REGION Network 26: fermer cv01 en 4k
   #_w1 := "EtatMode4k" AND NOT "CV01_ManAuto";
   IF #_w1 THEN
       "unscal_ret_val" := UNSCALE(IN := 0.0,
                               HI_LIM := 100.0,
                               LO_LIM := 0.0,
                               BIPOLAR := "always_0",
                               OUT => "CMD_CV_01");
       "PLC_to_Epics".CV01.sSetVAuto := 0.0;
   END_IF;
END_REGION

REGION Network 27: 2K mode - close CV02 after precooling the 2K line
   #_w1 := "EtatMode2K" AND (#S8step > 4);
   IF #_w1 THEN
       "unscal_ret_val_1" := UNSCALE(IN := 0.0,
                               HI_LIM := 100.0,
                               LO_LIM := 0.0,
                               BIPOLAR := "always_0",
                               OUT => "CMD_CV_02");
       "PLC_to_Epics".CV02.sSetVAuto := 0.0;
   END_IF;
END_REGION

REGION Network 28: Init 2K mode
   #_w1 := "EtatMode2K" AND NOT "2KModeStart_mem";   // rising edge of "EtatMode2K"
   "2KModeStart_mem" := "EtatMode2K";
   IF #_w1 THEN
       #S8step := 4;
       "unscal_ret_val" := UNSCALE(IN := "S8_parameters".CV01_Init,
                               HI_LIM := 100.0,
                               LO_LIM := 0.0,
                               BIPOLAR := "always_0",
                               OUT => "CMD_CV_01");
       "PLC_to_Epics".CV01.sSetVAuto := "S8_parameters".CV01_Init;
   END_IF;
END_REGION

REGION Network 29: 2K mode - precooling (step4)
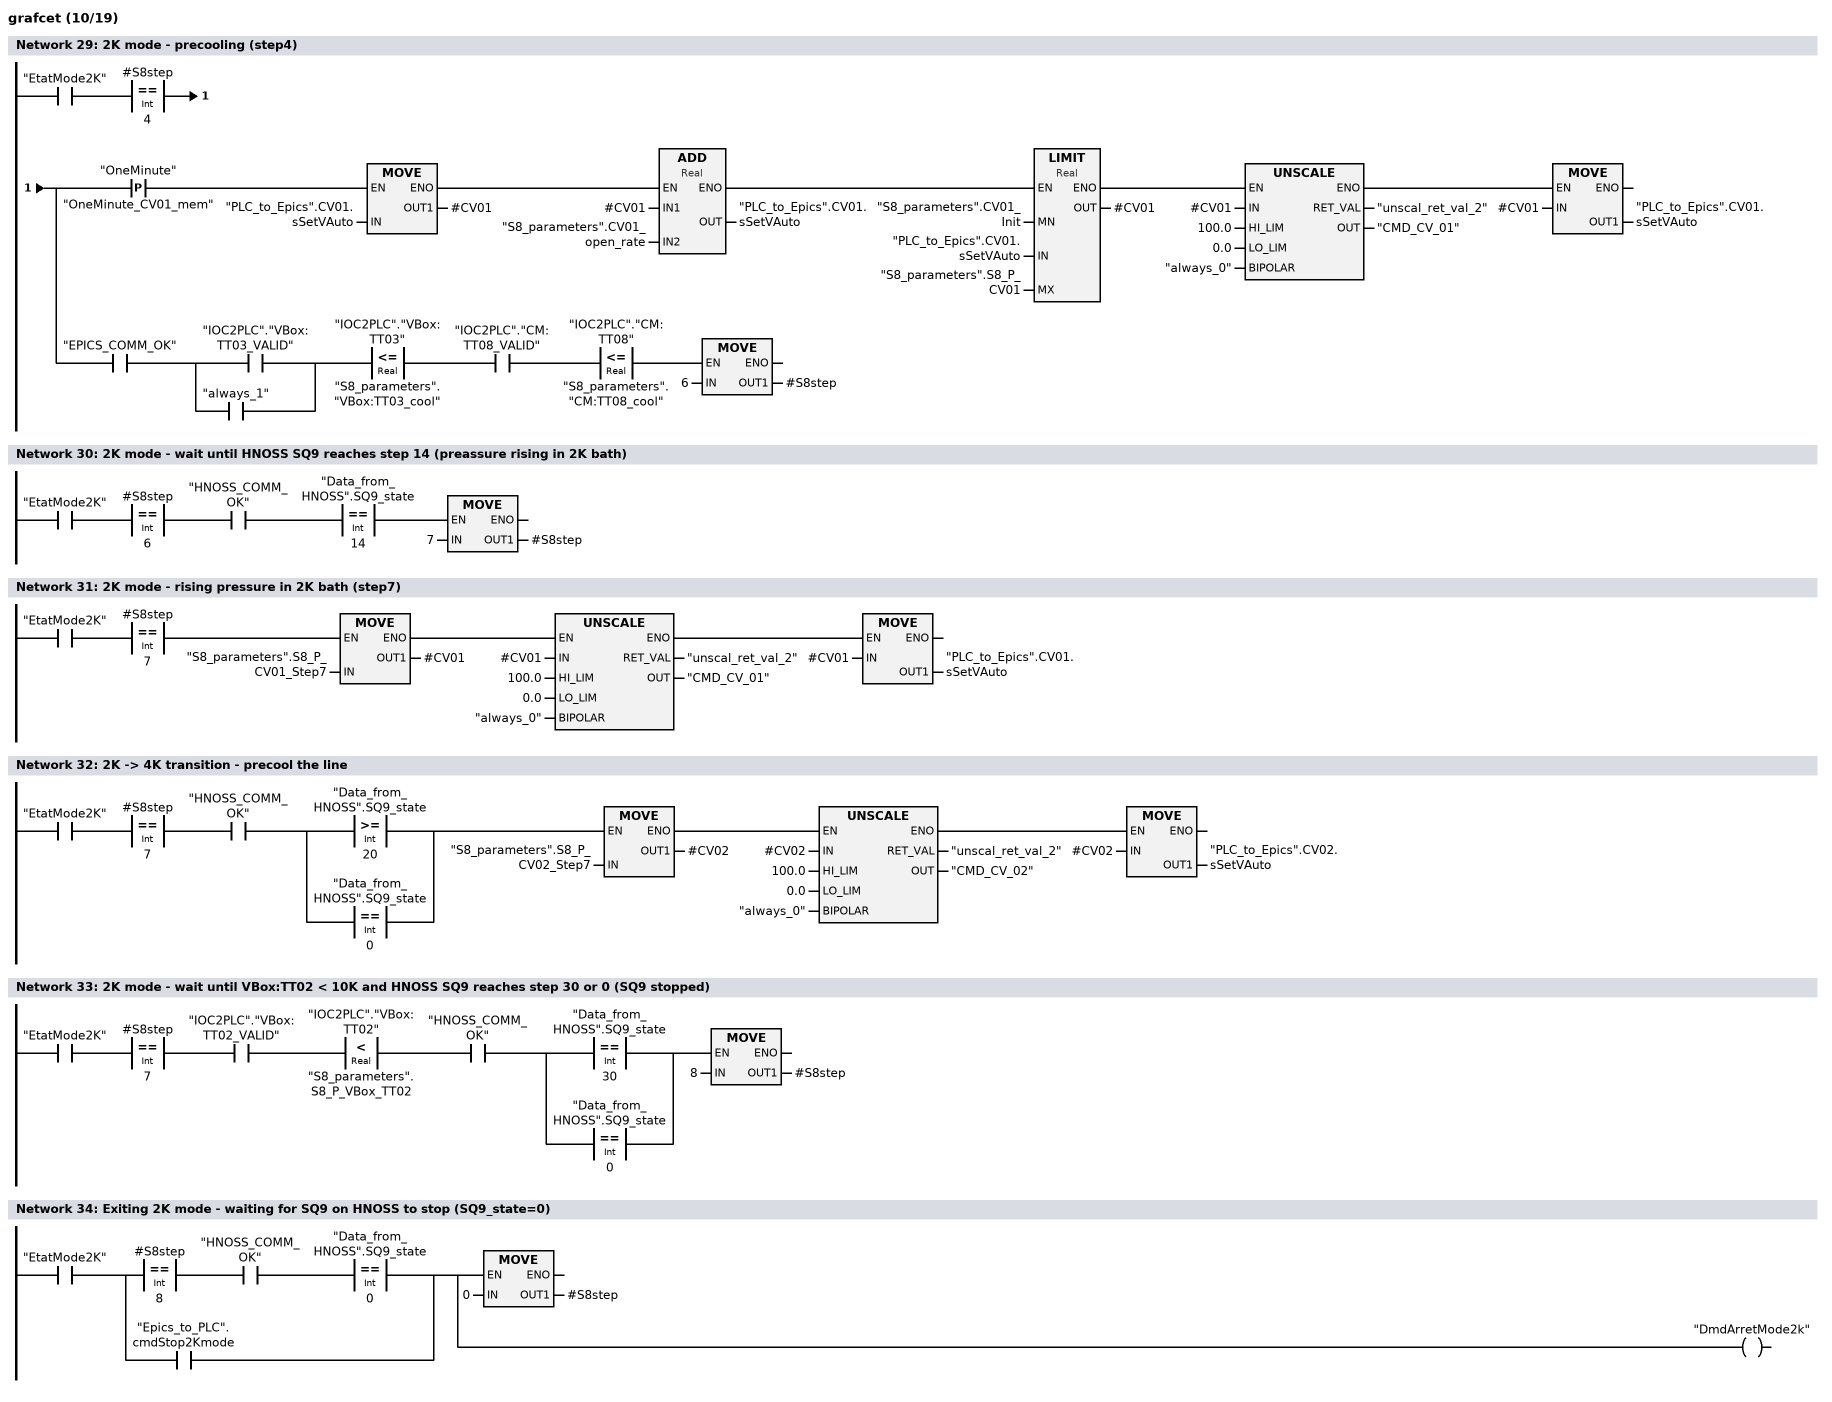
   // ENO of a box is taken as its EN; it also drops when the box reports an error
   #_w1 := "EtatMode2K" AND (#S8step = 4);
   #_w2 := #_w1 AND "OneMinute" AND NOT "OneMinute_CV01_mem";   // rising edge of "OneMinute"
   "OneMinute_CV01_mem" := "OneMinute";
   IF #_w2 THEN
       #CV01 := "PLC_to_Epics".CV01.sSetVAuto;
       "PLC_to_Epics".CV01.sSetVAuto := #CV01 + "S8_parameters".CV01_open_rate;
       #CV01 := LIMIT(MN := "S8_parameters".CV01_Init, IN := "PLC_to_Epics".CV01.sSetVAuto, MX := "S8_parameters".S8_P_CV01);
       "unscal_ret_val_2" := UNSCALE(IN := #CV01,
                               HI_LIM := 100.0,
                               LO_LIM := 0.0,
                               BIPOLAR := "always_0",
                               OUT => "CMD_CV_01");
       "PLC_to_Epics".CV01.sSetVAuto := #CV01;
   END_IF;
   IF #_w1 AND "EPICS_COMM_OK" AND ("IOC2PLC"."VBox:TT03_VALID" OR "always_1") AND ("IOC2PLC"."VBox:TT03" <= "S8_parameters"."VBox:TT03_cool") AND "IOC2PLC"."CM:TT08_VALID" AND ("IOC2PLC"."CM:TT08" <= "S8_parameters"."CM:TT08_cool") THEN
       #S8step := 6;
   END_IF;
END_REGION

REGION Network 30: 2K mode - wait until HNOSS SQ9 reaches step 14 (preassure rising in 2K bath)
   RUNG wire#powerrail
      Contact( "EtatMode2K" )
      { S7_Templates := "SrcType := Int" } EQ_Contact(in1 := #S8step, in2 := 6)
      Contact( "HNOSS_COMM_OK" )
      { S7_Templates := "SrcType := Int" } EQ_Contact(in1 := "Data_from_HNOSS".SQ9_state, in2 := 14)
      { S7_GenerateENO := "TRUE" } Move(in := 7, out1 => #S8step)
   END_RUNG
   // the same network as SCL:
   IF "EtatMode2K" AND (#S8step = 6) AND "HNOSS_COMM_OK" AND ("Data_from_HNOSS".SQ9_state = 14) THEN
       #S8step := 7;
   END_IF;
END_REGION

REGION Network 31: 2K mode - rising pressure in 2K bath (step7)
   // ENO of a box is taken as its EN; it also drops when the box reports an error
   IF "EtatMode2K" AND (#S8step = 7) THEN #CV01 := "S8_parameters".S8_P_CV01_Step7; END_IF;
   #_w1 := "EtatMode2K" AND (#S8step = 7);
   IF #_w1 THEN
       "unscal_ret_val_2" := UNSCALE(IN := #CV01,
                               HI_LIM := 100.0,
                               LO_LIM := 0.0,
                               BIPOLAR := "always_0",
                               OUT => "CMD_CV_01");
       "PLC_to_Epics".CV01.sSetVAuto := #CV01;
   END_IF;
END_REGION

REGION Network 32: 2K -> 4K transition - precool the line
   // ENO of a box is taken as its EN; it also drops when the box reports an error
   IF "EtatMode2K" AND (#S8step = 7) AND "HNOSS_COMM_OK" AND (("Data_from_HNOSS".SQ9_state >= 20) OR ("Data_from_HNOSS".SQ9_state = 0)) THEN
       #CV02 := "S8_parameters".S8_P_CV02_Step7;
   END_IF;
   #_w1 := "EtatMode2K" AND (#S8step = 7) AND "HNOSS_COMM_OK" AND (("Data_from_HNOSS".SQ9_state >= 20) OR ("Data_from_HNOSS".SQ9_state = 0));
   IF #_w1 THEN
       "unscal_ret_val_2" := UNSCALE(IN := #CV02,
                               HI_LIM := 100.0,
                               LO_LIM := 0.0,
                               BIPOLAR := "always_0",
                               OUT => "CMD_CV_02");
       "PLC_to_Epics".CV02.sSetVAuto := #CV02;
   END_IF;
END_REGION

REGION Network 33: 2K mode - wait until VBox:TT02 < 10K and HNOSS SQ9 reaches step 30 or 0 (SQ9 stopped)
   RUNG wire#powerrail
      Contact( "EtatMode2K" )
      { S7_Templates := "SrcType := Int" } EQ_Contact(in1 := #S8step, in2 := 7)
      Contact( "IOC2PLC"."VBox:TT02_VALID" )
      { S7_Templates := "SrcType := Real" } LT_Contact(in1 := "IOC2PLC"."VBox:TT02", in2 := "S8_parameters".S8_P_VBox_TT02)
      Contact( "HNOSS_COMM_OK" )
      wire#w1
      { S7_Templates := "SrcType := Int" } EQ_Contact(in1 := "Data_from_HNOSS".SQ9_state, in2 := 30)
      wire#w2
      { S7_GenerateENO := "TRUE" } Move(in := 8, out1 => #S8step)
   END_RUNG
   RUNG wire#w1
      { S7_Templates := "SrcType := Int" } EQ_Contact(in1 := "Data_from_HNOSS".SQ9_state, in2 := 0)
   END_RUNG wire#w2
   // the same network as SCL:
   IF "EtatMode2K" AND (#S8step = 7) AND "IOC2PLC"."VBox:TT02_VALID" AND ("IOC2PLC"."VBox:TT02" < "S8_parameters".S8_P_VBox_TT02) AND "HNOSS_COMM_OK" AND (("Data_from_HNOSS".SQ9_state = 30) OR ("Data_from_HNOSS".SQ9_state = 0)) THEN
       #S8step := 8;
   END_IF;
END_REGION

REGION Network 34: Exiting 2K mode - waiting for SQ9 on HNOSS to stop (SQ9_state=0)
   RUNG wire#powerrail
      Contact( "EtatMode2K" )
      wire#w1
      { S7_Templates := "SrcType := Int" } EQ_Contact(in1 := #S8step, in2 := 8)
      Contact( "HNOSS_COMM_OK" )
      { S7_Templates := "SrcType := Int" } EQ_Contact(in1 := "Data_from_HNOSS".SQ9_state, in2 := 0)
      wire#w2
      { S7_GenerateENO := "TRUE" } Move(in := 0, out1 => #S8step)
   END_RUNG
   RUNG wire#w1
      Contact( "Epics_to_PLC".cmdStop2Kmode )
   END_RUNG wire#w2
   RUNG wire#w2
      Coil( "DmdArretMode2k" )
   END_RUNG
   // the same network as SCL:
   #_w1 := "EtatMode2K" AND (((#S8step = 8) AND "HNOSS_COMM_OK" AND ("Data_from_HNOSS".SQ9_state = 0)) OR "Epics_to_PLC".cmdStop2Kmode);
   IF #_w1 THEN #S8step := 0; END_IF;
   "DmdArretMode2k" := #_w1;
END_REGION

REGION Network 35: Config vannes mode standby
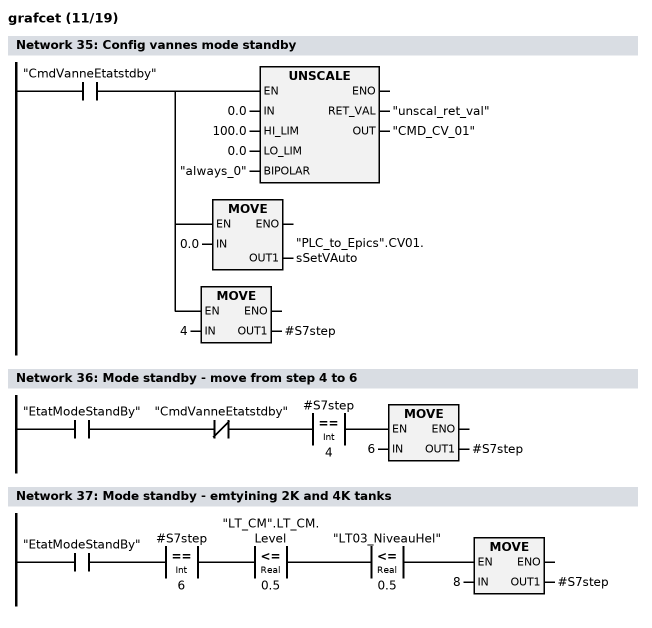
   #_w1 := "CmdVanneEtatstdby";
   IF #_w1 THEN
       "unscal_ret_val" := UNSCALE(IN := 0.0,
                               HI_LIM := 100.0,
                               LO_LIM := 0.0,
                               BIPOLAR := "always_0",
                               OUT => "CMD_CV_01");
       "PLC_to_Epics".CV01.sSetVAuto := 0.0;
       #S7step := 4;
   END_IF;
END_REGION

REGION Network 36: Mode standby - move from step 4 to 6
   RUNG wire#powerrail
      Contact( "EtatModeStandBy" )
      I_Contact( "CmdVanneEtatstdby" )
      { S7_Templates := "SrcType := Int" } EQ_Contact(in1 := #S7step, in2 := 4)
      { S7_GenerateENO := "TRUE" } Move(in := 6, out1 => #S7step)
   END_RUNG
   // the same network as SCL:
   IF "EtatModeStandBy" AND NOT "CmdVanneEtatstdby" AND (#S7step = 4) THEN #S7step := 6; END_IF;
END_REGION

REGION Network 37: Mode standby - emtyining 2K and 4K tanks
   RUNG wire#powerrail
      Contact( "EtatModeStandBy" )
      { S7_Templates := "SrcType := Int" } EQ_Contact(in1 := #S7step, in2 := 6)
      { S7_Templates := "SrcType := Real" } LE_Contact(in1 := "LT_CM".LT_CM.Level, in2 := 0.5)
      { S7_Templates := "SrcType := Real" } LE_Contact(in1 := "LT03_NiveauHel", in2 := 0.5)
      { S7_GenerateENO := "TRUE" } Move(in := 8, out1 => #S7step)
   END_RUNG
   // the same network as SCL:
   IF "EtatModeStandBy" AND (#S7step = 6) AND ("LT_CM".LT_CM.Level <= 0.5) AND ("LT03_NiveauHel" <= 0.5) THEN
       #S7step := 8;
   END_IF;
END_REGION

REGION Network 38: Mode standby - warming up (step8) and cooling (step10)
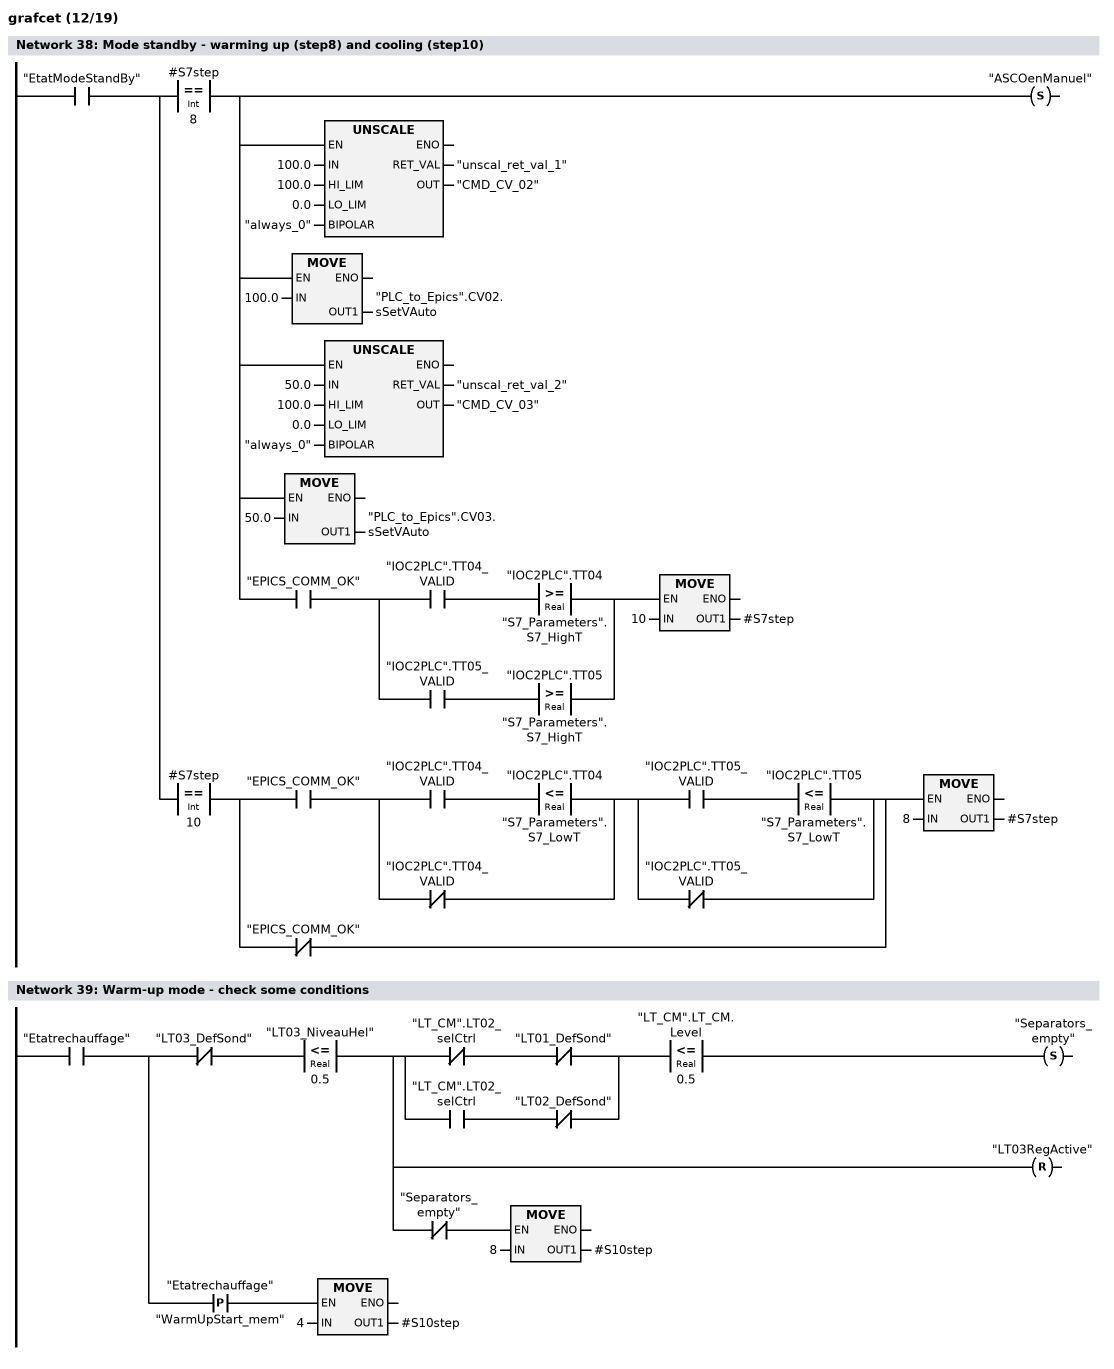
   #_w1 := "EtatModeStandBy" AND (#S7step = 8);
   IF #_w1 THEN "ASCOenManuel" := TRUE; END_IF;
   #_w2 := "EtatModeStandBy";
   IF #_w1 THEN
       "unscal_ret_val_1" := UNSCALE(IN := 100.0,
                               HI_LIM := 100.0,
                               LO_LIM := 0.0,
                               BIPOLAR := "always_0",
                               OUT => "CMD_CV_02");
       "PLC_to_Epics".CV02.sSetVAuto := 100.0;
       "unscal_ret_val_2" := UNSCALE(IN := 50.0,
                               HI_LIM := 100.0,
                               LO_LIM := 0.0,
                               BIPOLAR := "always_0",
                               OUT => "CMD_CV_03");
       "PLC_to_Epics".CV03.sSetVAuto := 50.0;
   END_IF;
   IF #_w1 AND "EPICS_COMM_OK" AND (("IOC2PLC".TT04_VALID AND ("IOC2PLC".TT04 >= "S7_Parameters".S7_HighT)) OR ("IOC2PLC".TT05_VALID AND ("IOC2PLC".TT05 >= "S7_Parameters".S7_HighT))) THEN
       #S7step := 10;
   END_IF;
   IF #_w2 AND (#S7step = 10) AND (("EPICS_COMM_OK" AND (("IOC2PLC".TT04_VALID AND ("IOC2PLC".TT04 <= "S7_Parameters".S7_LowT)) OR NOT "IOC2PLC".TT04_VALID) AND (("IOC2PLC".TT05_VALID AND ("IOC2PLC".TT05 <= "S7_Parameters".S7_LowT)) OR NOT "IOC2PLC".TT05_VALID)) OR NOT "EPICS_COMM_OK") THEN
       #S7step := 8;
   END_IF;
END_REGION

REGION Network 39: Warm-up mode - check some conditions
   RUNG wire#powerrail
      Contact( "Etatrechauffage" )
      wire#w1
      I_Contact( "LT03_DefSond" )
      { S7_Templates := "SrcType := Real" } LE_Contact(in1 := "LT03_NiveauHel", in2 := 0.5)
      wire#w2
      I_Contact( "LT_CM".LT02_selCtrl )
      I_Contact( "LT01_DefSond" )
      wire#w3
      { S7_Templates := "SrcType := Real" } LE_Contact(in1 := "LT_CM".LT_CM.Level, in2 := 0.5)
      S_Coil( "Separators_empty" )
   END_RUNG
   RUNG wire#w2
      Contact( "LT_CM".LT02_selCtrl )
      I_Contact( "LT02_DefSond" )
   END_RUNG wire#w3
   RUNG wire#w2
      R_Coil( "LT03RegActive" )
   END_RUNG
   RUNG wire#w2
      I_Contact( "Separators_empty" )
      { S7_GenerateENO := "TRUE" } Move(in := 8, out1 => #S10step)
   END_RUNG
   RUNG wire#w1
      P_Contact(operand := "Etatrechauffage", bit := "WarmUpStart_mem")
      { S7_GenerateENO := "TRUE" } Move(in := 4, out1 => #S10step)
   END_RUNG
   // the same network as SCL:
   #_w1 := "Etatrechauffage" AND NOT "LT03_DefSond" AND ("LT03_NiveauHel" <= 0.5);
   IF #_w1 AND ((NOT "LT_CM".LT02_selCtrl AND NOT "LT01_DefSond") OR ("LT_CM".LT02_selCtrl AND NOT "LT02_DefSond")) AND ("LT_CM".LT_CM.Level <= 0.5) THEN
       "Separators_empty" := TRUE;
   END_IF;
   IF #_w1 THEN "LT03RegActive" := FALSE; END_IF;
   IF #_w1 AND NOT "Separators_empty" THEN #S10step := 8; END_IF;
   #_w2 := "Etatrechauffage" AND "Etatrechauffage" AND NOT "WarmUpStart_mem";   // rising edge of "Etatrechauffage"
   "WarmUpStart_mem" := "Etatrechauffage";
   IF #_w2 THEN #S10step := 4; END_IF;
END_REGION

REGION Network 40: Warm-up: set-up the settings of CV01-CV04
   // Set-up the settings depending on the LHe levels in the phase separators
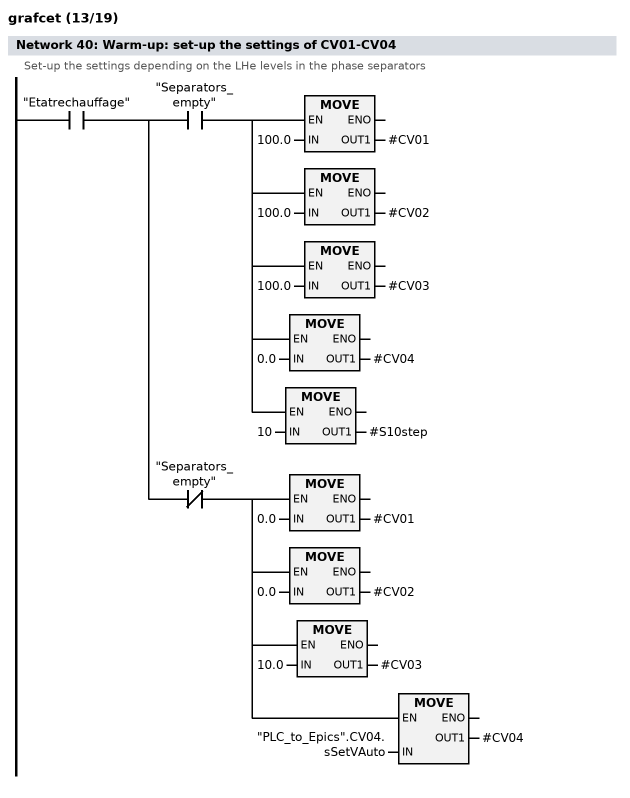
   RUNG wire#powerrail
      Contact( "Etatrechauffage" )
      wire#w1
      Contact( "Separators_empty" )
      wire#w2
      { S7_GenerateENO := "TRUE" } Move(in := 100.0, out1 => #CV01)
   END_RUNG
   RUNG wire#w2
      { S7_GenerateENO := "TRUE" } Move(in := 100.0, out1 => #CV02)
   END_RUNG
   RUNG wire#w2
      { S7_GenerateENO := "TRUE" } Move(in := 100.0, out1 => #CV03)
   END_RUNG
   RUNG wire#w2
      { S7_GenerateENO := "TRUE" } Move(in := 0.0, out1 => #CV04)
   END_RUNG
   RUNG wire#w2
      { S7_GenerateENO := "TRUE" } Move(in := 10, out1 => #S10step)
   END_RUNG
   RUNG wire#w1
      I_Contact( "Separators_empty" )
      wire#w3
      { S7_GenerateENO := "TRUE" } Move(in := 0.0, out1 => #CV01)
   END_RUNG
   RUNG wire#w3
      { S7_GenerateENO := "TRUE" } Move(in := 0.0, out1 => #CV02)
   END_RUNG
   RUNG wire#w3
      { S7_GenerateENO := "TRUE" } Move(in := 10.0, out1 => #CV03)
   END_RUNG
   RUNG wire#w3
      { S7_GenerateENO := "TRUE" } Move(in := "PLC_to_Epics".CV04.sSetVAuto, out1 => #CV04)
   END_RUNG
   // the same network as SCL:
   IF "Etatrechauffage" AND "Separators_empty" THEN
       #CV01 := 100.0;
       #CV02 := 100.0;
       #CV03 := 100.0;
       #CV04 := 0.0;
       #S10step := 10;
   END_IF;
   IF "Etatrechauffage" AND NOT "Separators_empty" THEN
       #CV01 := 0.0;
       #CV02 := 0.0;
       #CV03 := 10.0;
       #CV04 := "PLC_to_Epics".CV04.sSetVAuto;
   END_IF;
END_REGION

REGION Network 41: Mode Rechauffage
   // The heaters are handled in Manage_HEATERS
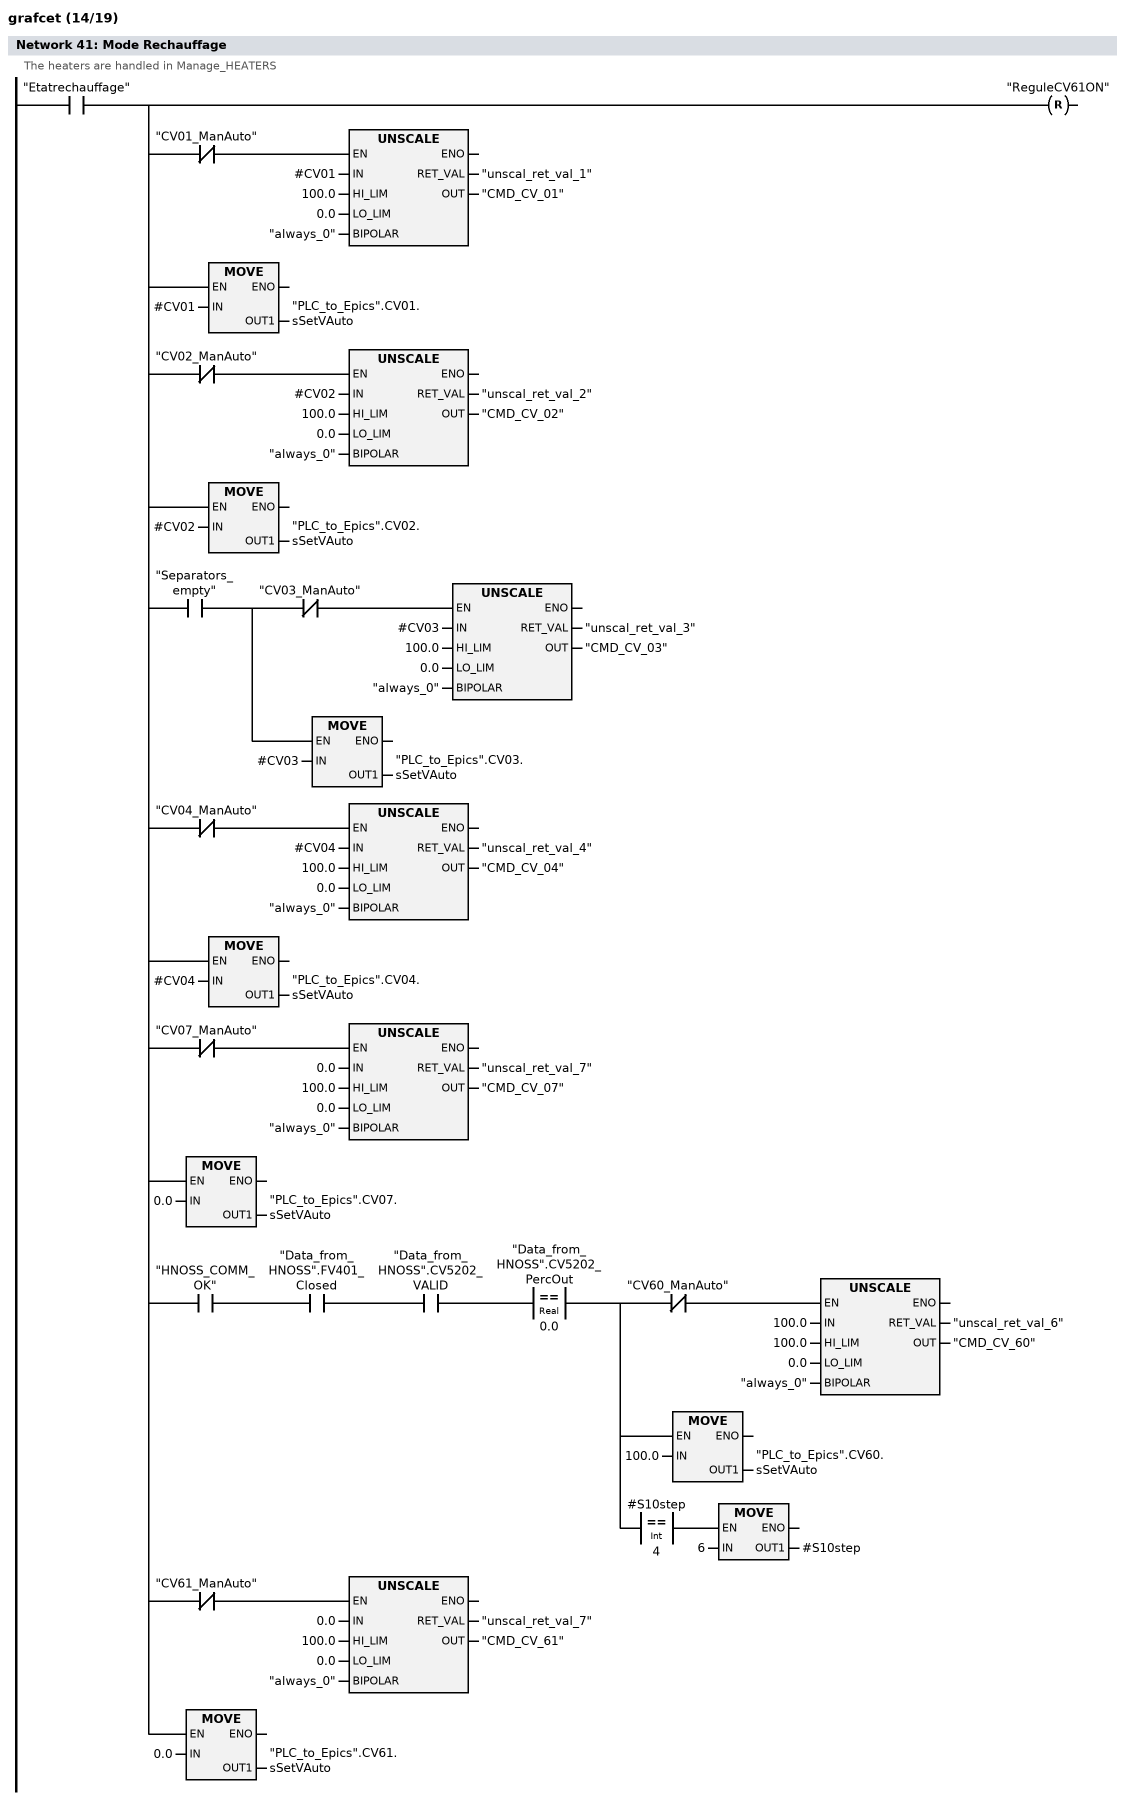
   IF "Etatrechauffage" THEN "ReguleCV61ON" := FALSE; END_IF;
   #_w1 := "Etatrechauffage";
   IF "Etatrechauffage" AND NOT "CV01_ManAuto" THEN
       "unscal_ret_val_1" := UNSCALE(IN := #CV01,
                               HI_LIM := 100.0,
                               LO_LIM := 0.0,
                               BIPOLAR := "always_0",
                               OUT => "CMD_CV_01");
   END_IF;
   IF #_w1 THEN "PLC_to_Epics".CV01.sSetVAuto := #CV01; END_IF;
   IF #_w1 AND NOT "CV02_ManAuto" THEN
       "unscal_ret_val_2" := UNSCALE(IN := #CV02,
                               HI_LIM := 100.0,
                               LO_LIM := 0.0,
                               BIPOLAR := "always_0",
                               OUT => "CMD_CV_02");
   END_IF;
   IF #_w1 THEN "PLC_to_Epics".CV02.sSetVAuto := #CV02; END_IF;
   #_w2 := #_w1 AND "Separators_empty";
   IF #_w2 AND NOT "CV03_ManAuto" THEN
       "unscal_ret_val_3" := UNSCALE(IN := #CV03,
                               HI_LIM := 100.0,
                               LO_LIM := 0.0,
                               BIPOLAR := "always_0",
                               OUT => "CMD_CV_03");
   END_IF;
   IF #_w2 THEN "PLC_to_Epics".CV03.sSetVAuto := #CV03; END_IF;
   IF #_w1 AND NOT "CV04_ManAuto" THEN
       "unscal_ret_val_4" := UNSCALE(IN := #CV04,
                               HI_LIM := 100.0,
                               LO_LIM := 0.0,
                               BIPOLAR := "always_0",
                               OUT => "CMD_CV_04");
   END_IF;
   IF #_w1 THEN "PLC_to_Epics".CV04.sSetVAuto := #CV04; END_IF;
   IF #_w1 AND NOT "CV07_ManAuto" THEN
       "unscal_ret_val_7" := UNSCALE(IN := 0.0,
                               HI_LIM := 100.0,
                               LO_LIM := 0.0,
                               BIPOLAR := "always_0",
                               OUT => "CMD_CV_07");
   END_IF;
   IF #_w1 THEN "PLC_to_Epics".CV07.sSetVAuto := 0.0; END_IF;
   #_w3 := #_w1 AND "HNOSS_COMM_OK" AND "Data_from_HNOSS".FV401_Closed AND "Data_from_HNOSS".CV5202_VALID AND ("Data_from_HNOSS".CV5202_PercOut = 0.0);
   IF #_w3 AND NOT "CV60_ManAuto" THEN
       "unscal_ret_val_6" := UNSCALE(IN := 100.0,
                               HI_LIM := 100.0,
                               LO_LIM := 0.0,
                               BIPOLAR := "always_0",
                               OUT => "CMD_CV_60");
   END_IF;
   IF #_w3 THEN "PLC_to_Epics".CV60.sSetVAuto := 100.0; END_IF;
   IF #_w3 AND (#S10step = 4) THEN #S10step := 6; END_IF;
   IF #_w1 AND NOT "CV61_ManAuto" THEN
       "unscal_ret_val_7" := UNSCALE(IN := 0.0,
                               HI_LIM := 100.0,
                               LO_LIM := 0.0,
                               BIPOLAR := "always_0",
                               OUT => "CMD_CV_61");
   END_IF;
   IF #_w1 THEN "PLC_to_Epics".CV61.sSetVAuto := 0.0; END_IF;
END_REGION

REGION Network 42: Mode manuel ASCO
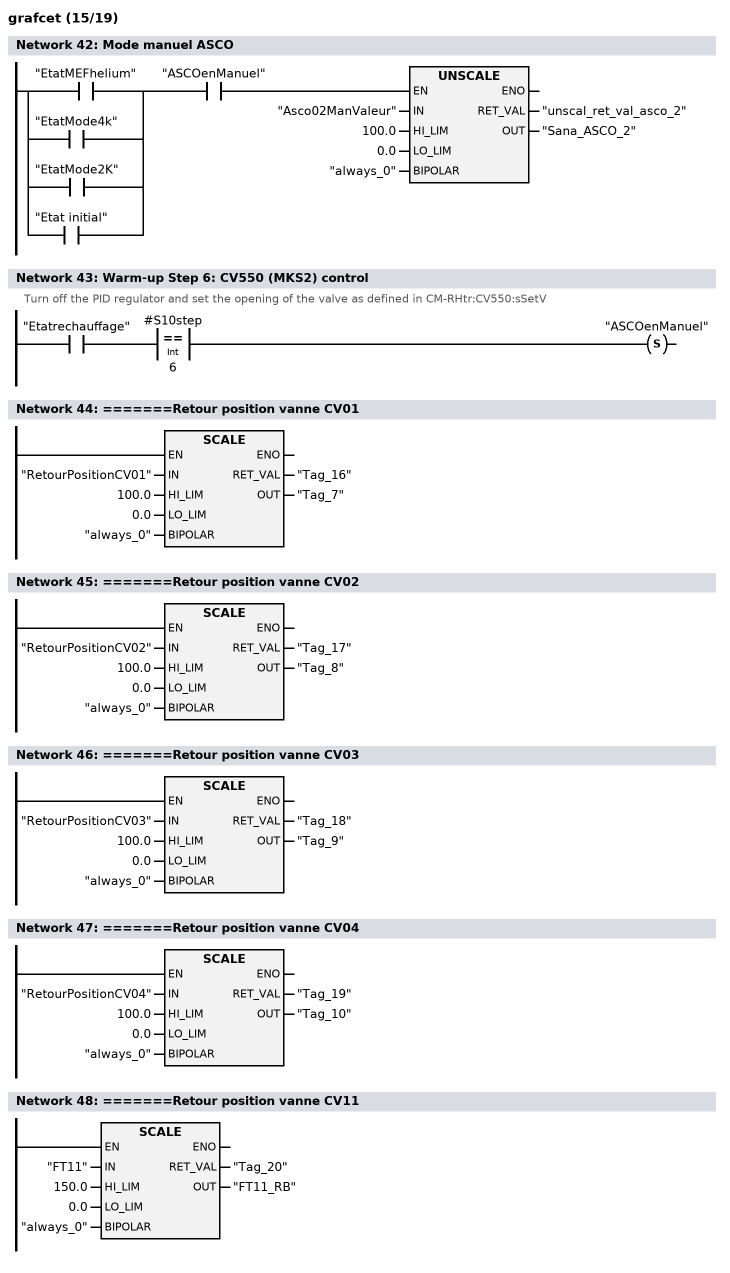
   IF ("EtatMEFhelium" OR "EtatMode4k" OR "EtatMode2K" OR "Etat initial") AND "ASCOenManuel" THEN
       "unscal_ret_val_asco_2" := UNSCALE(in := "Asco02ManValeur",
                               hi_lim := 100.0,
                               lo_lim := 0.0,
                               bipolar := "always_0",
                               out => "Sana_ASCO_2");
   END_IF;
END_REGION

REGION Network 43: Warm-up Step 6: CV550 (MKS2) control
   // Turn off the PID regulator and set the opening of the valve as defined in CM-RHtr:CV550:sSetV
   RUNG wire#powerrail
      Contact( "Etatrechauffage" )
      { S7_Templates := "SrcType := Int" } EQ_Contact(in1 := #S10step, in2 := 6)
      S_Coil( "ASCOenManuel" )
   END_RUNG
   // the same network as SCL:
   IF "Etatrechauffage" AND (#S10step = 6) THEN "ASCOenManuel" := TRUE; END_IF;
END_REGION

REGION Network 44: =======Retour position vanne CV01
   "Tag_16" := SCALE(in := "RetourPositionCV01",
                     hi_lim := 100.0,
                     lo_lim := 0.0,
                     bipolar := "always_0",
                     out => "Tag_7");
END_REGION

REGION Network 45: =======Retour position vanne CV02
   "Tag_17" := SCALE(in := "RetourPositionCV02",
                     hi_lim := 100.0,
                     lo_lim := 0.0,
                     bipolar := "always_0",
                     out => "Tag_8");
END_REGION

REGION Network 46: =======Retour position vanne CV03
   "Tag_18" := SCALE(in := "RetourPositionCV03",
                     hi_lim := 100.0,
                     lo_lim := 0.0,
                     bipolar := "always_0",
                     out => "Tag_9");
END_REGION

REGION Network 47: =======Retour position vanne CV04
   "Tag_19" := SCALE(in := "RetourPositionCV04",
                     hi_lim := 100.0,
                     lo_lim := 0.0,
                     bipolar := "always_0",
                     out => "Tag_10");
END_REGION

REGION Network 48: =======Retour position vanne CV11
   "Tag_20" := SCALE(IN := "FT11", HI_LIM := 150.0, LO_LIM := 0.0, BIPOLAR := "always_0", OUT => "FT11_RB");
END_REGION

REGION Network 49: =======Retour position vanne CV21
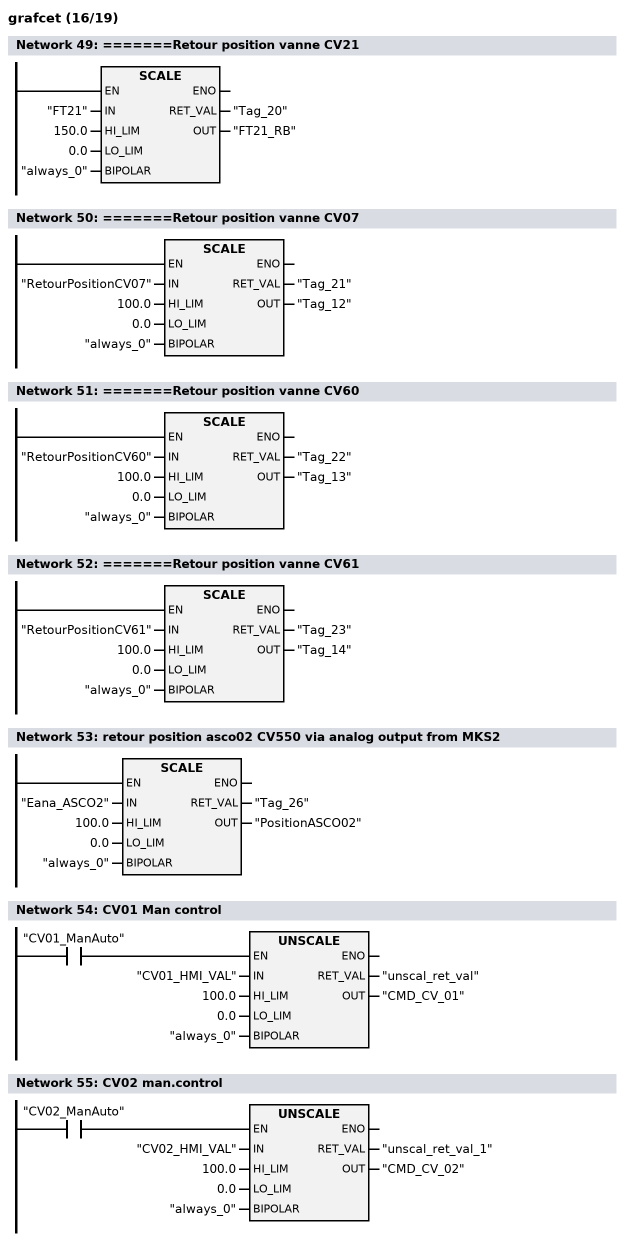
   "Tag_20" := SCALE(IN := "FT21", HI_LIM := 150.0, LO_LIM := 0.0, BIPOLAR := "always_0", OUT => "FT21_RB");
END_REGION

REGION Network 50: =======Retour position vanne CV07
   "Tag_21" := SCALE(in := "RetourPositionCV07",
                     hi_lim := 100.0,
                     lo_lim := 0.0,
                     bipolar := "always_0",
                     out => "Tag_12");
END_REGION

REGION Network 51: =======Retour position vanne CV60
   "Tag_22" := SCALE(in := "RetourPositionCV60",
                     hi_lim := 100.0,
                     lo_lim := 0.0,
                     bipolar := "always_0",
                     out => "Tag_13");
END_REGION

REGION Network 52: =======Retour position vanne CV61
   "Tag_23" := SCALE(in := "RetourPositionCV61",
                     hi_lim := 100.0,
                     lo_lim := 0.0,
                     bipolar := "always_0",
                     out => "Tag_14");
END_REGION

REGION Network 53: retour position asco02 CV550 via analog output from MKS2
   "Tag_26" := SCALE(in := "Eana_ASCO2",
                     hi_lim := 100.0,
                     lo_lim := 0.0,
                     bipolar := "always_0",
                     out => "PositionASCO02");
END_REGION

REGION Network 54: CV01 Man control
   IF "CV01_ManAuto" THEN
       "unscal_ret_val" := UNSCALE(in := "CV01_HMI_VAL",
                               hi_lim := 100.0,
                               lo_lim := 0.0,
                               bipolar := "always_0",
                               out => "CMD_CV_01");
   END_IF;
END_REGION

REGION Network 55: CV02 man.control
   IF "CV02_ManAuto" THEN
       "unscal_ret_val_1" := UNSCALE(in := "CV02_HMI_VAL",
                               hi_lim := 100.0,
                               lo_lim := 0.0,
                               bipolar := "always_0",
                               out => "CMD_CV_02");
   END_IF;
END_REGION

REGION Network 56: CV03 manual control
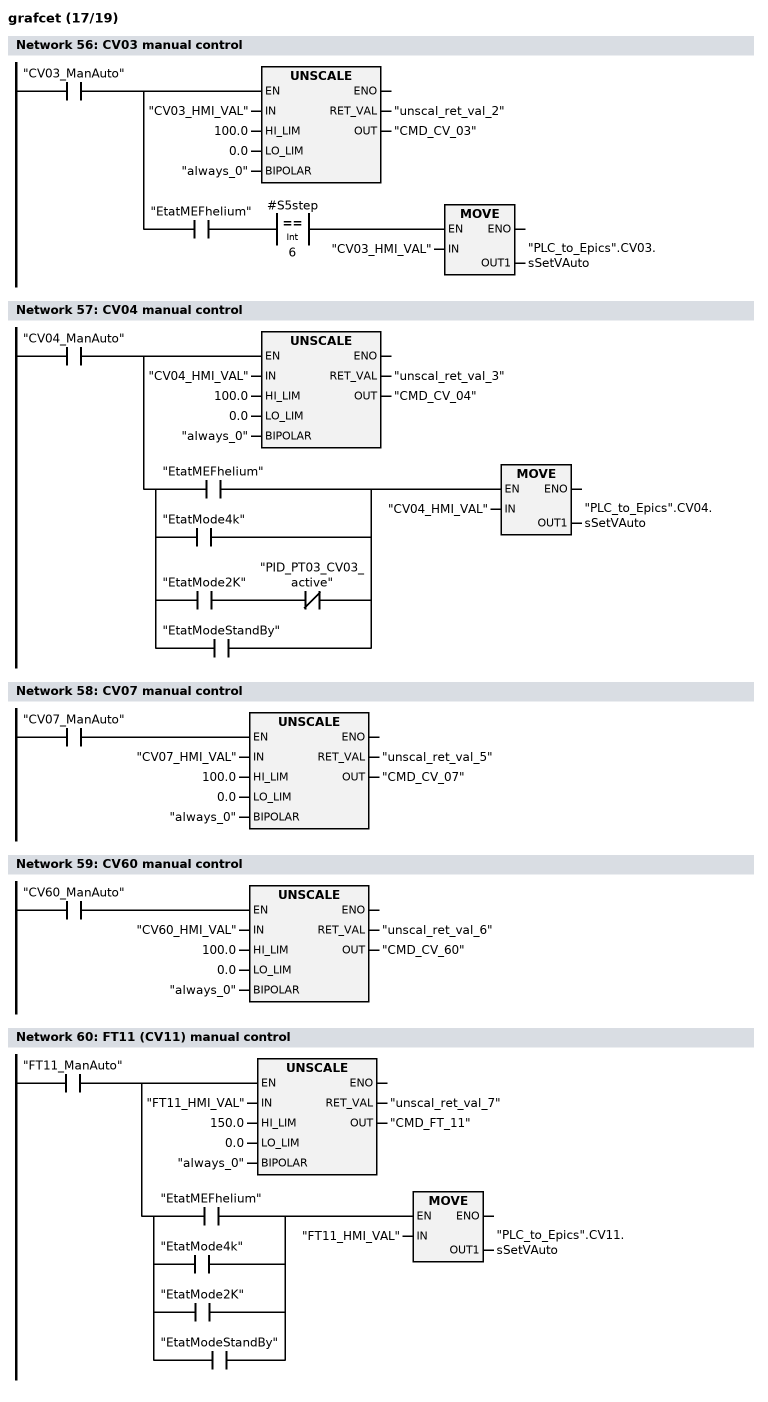
   #_w1 := "CV03_ManAuto";
   IF #_w1 THEN
       "unscal_ret_val_2" := UNSCALE(IN := "CV03_HMI_VAL",
                               HI_LIM := 100.0,
                               LO_LIM := 0.0,
                               BIPOLAR := "always_0",
                               OUT => "CMD_CV_03");
   END_IF;
   IF #_w1 AND "EtatMEFhelium" AND (#S5step = 6) THEN
       "PLC_to_Epics".CV03.sSetVAuto := "CV03_HMI_VAL";
   END_IF;
END_REGION

REGION Network 57: CV04 manual control
   #_w1 := "CV04_ManAuto";
   IF #_w1 THEN
       "unscal_ret_val_3" := UNSCALE(IN := "CV04_HMI_VAL",
                               HI_LIM := 100.0,
                               LO_LIM := 0.0,
                               BIPOLAR := "always_0",
                               OUT => "CMD_CV_04");
   END_IF;
   IF #_w1 AND ("EtatMEFhelium" OR "EtatMode4k" OR ("EtatMode2K" AND NOT "PID_PT03_CV03_active") OR "EtatModeStandBy") THEN
       "PLC_to_Epics".CV04.sSetVAuto := "CV04_HMI_VAL";
   END_IF;
END_REGION

REGION Network 58: CV07 manual control
   IF "CV07_ManAuto" THEN
       "unscal_ret_val_5" := UNSCALE(in := "CV07_HMI_VAL",
                               hi_lim := 100.0,
                               lo_lim := 0.0,
                               bipolar := "always_0",
                               out => "CMD_CV_07");
   END_IF;
END_REGION

REGION Network 59: CV60 manual control
   IF "CV60_ManAuto" THEN
       "unscal_ret_val_6" := UNSCALE(in := "CV60_HMI_VAL",
                               hi_lim := 100.0,
                               lo_lim := 0.0,
                               bipolar := "always_0",
                               out => "CMD_CV_60");
   END_IF;
END_REGION

REGION Network 60: FT11 (CV11) manual control
   #_w1 := "FT11_ManAuto";
   IF #_w1 THEN
       "unscal_ret_val_7" := UNSCALE(IN := "FT11_HMI_VAL",
                               HI_LIM := 150.0,
                               LO_LIM := 0.0,
                               BIPOLAR := "always_0",
                               OUT => "CMD_FT_11");
   END_IF;
   IF #_w1 AND ("EtatMEFhelium" OR "EtatMode4k" OR "EtatMode2K" OR "EtatModeStandBy") THEN
       "PLC_to_Epics".CV11.sSetVAuto := "FT11_HMI_VAL";
   END_IF;
END_REGION

REGION Network 61: FT21 (CV21) manual control
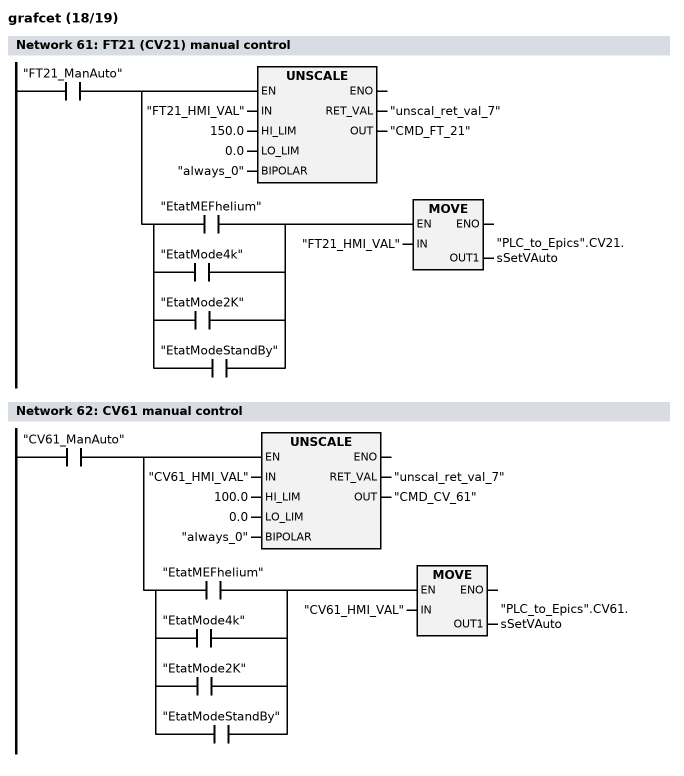
   #_w1 := "FT21_ManAuto";
   IF #_w1 THEN
       "unscal_ret_val_7" := UNSCALE(IN := "FT21_HMI_VAL",
                               HI_LIM := 150.0,
                               LO_LIM := 0.0,
                               BIPOLAR := "always_0",
                               OUT => "CMD_FT_21");
   END_IF;
   IF #_w1 AND ("EtatMEFhelium" OR "EtatMode4k" OR "EtatMode2K" OR "EtatModeStandBy") THEN
       "PLC_to_Epics".CV21.sSetVAuto := "FT21_HMI_VAL";
   END_IF;
END_REGION

REGION Network 62: CV61 manual control
   #_w1 := "CV61_ManAuto";
   IF #_w1 THEN
       "unscal_ret_val_7" := UNSCALE(IN := "CV61_HMI_VAL",
                               HI_LIM := 100.0,
                               LO_LIM := 0.0,
                               BIPOLAR := "always_0",
                               OUT => "CMD_CV_61");
   END_IF;
   IF #_w1 AND ("EtatMEFhelium" OR "EtatMode4k" OR "EtatMode2K" OR "EtatModeStandBy") THEN
       "PLC_to_Epics".CV61.sSetVAuto := "CV61_HMI_VAL";
   END_IF;
END_REGION

REGION Network 63: Graph
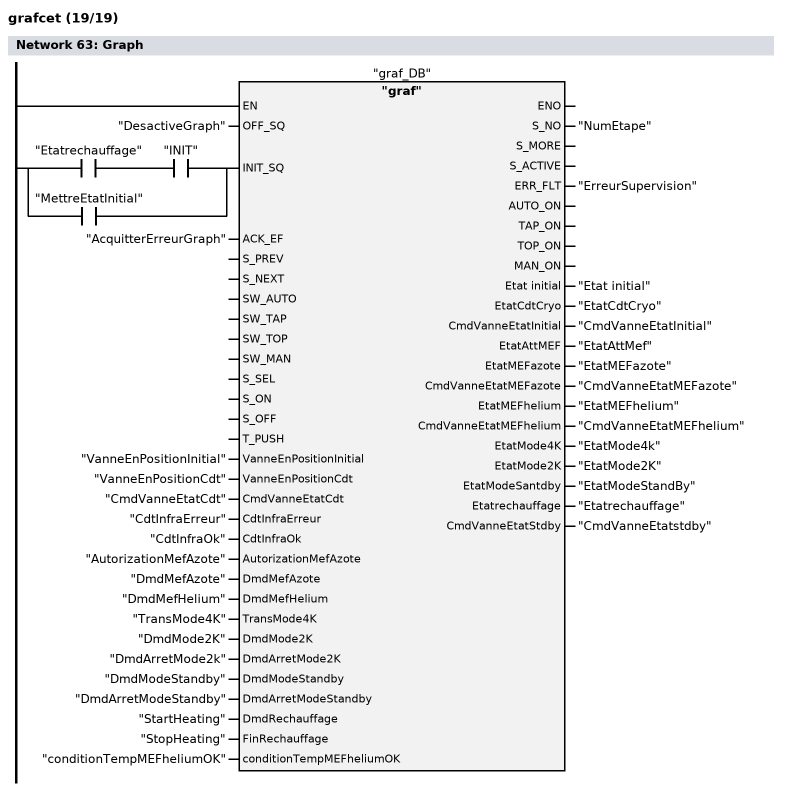
   "graf_DB"(OFF_SQ := "DesactiveGraph",   // "graf"
             INIT_SQ := "MettreEtatInitial" OR ("Etatrechauffage" AND "INIT"),
             ACK_EF := "AcquitterErreurGraph",
             VanneEnPositionInitial := "VanneEnPositionInitial",
             VanneEnPositionCdt := "VanneEnPositionCdt",
             CmdVanneEtatCdt := "CmdVanneEtatCdt",
             CdtInfraErreur := "CdtInfraErreur",
             CdtInfraOk := "CdtInfraOk",
             AutorizationMefAzote := "AutorizationMefAzote",
             DmdMefAzote := "DmdMefAzote",
             DmdMefHelium := "DmdMefHelium",
             TransMode4K := "TransMode4K",
             DmdMode2K := "DmdMode2K",
             DmdArretMode2K := "DmdArretMode2k",
             DmdModeStandby := "DmdModeStandby",
             DmdArretModeStandby := "DmdArretModeStandby",
             DmdRechauffage := "StartHeating",
             FinRechauffage := "StopHeating",
             conditionTempMEFheliumOK := "conditionTempMEFheliumOK",
             S_NO => "NumEtape",
             ERR_FLT => "ErreurSupervision",
             "Etat initial" => "Etat initial",
             EtatCdtCryo => "EtatCdtCryo",
             CmdVanneEtatInitial => "CmdVanneEtatInitial",
             EtatAttMEF => "EtatAttMef",
             EtatMEFazote => "EtatMEFazote",
             CmdVanneEtatMEFazote => "CmdVanneEtatMEFazote",
             EtatMEFhelium => "EtatMEFhelium",
             CmdVanneEtatMEFhelium => "CmdVanneEtatMEFhelium",
             EtatMode4K => "EtatMode4k",
             EtatMode2K => "EtatMode2K",
             EtatModeSantdby => "EtatModeStandBy",
             Etatrechauffage => "Etatrechauffage",
             CmdVanneEtatStdby => "CmdVanneEtatstdby");
END_REGION

REGION Network 64 (STL): Copy step number to HNOSS
         L     #S4step;
         T     "Data_to_HNOSS".S4step;
         L     #S5step;
         T     "Data_to_HNOSS".S5step;
         L     #S6step;
         T     "Data_to_HNOSS".S6step;
         L     #S7step;
         T     "Data_to_HNOSS".S7step;
         L     #S8step;
         T     "Data_to_HNOSS".S8step;
         L     #S9step;
         T     "Data_to_HNOSS".S9step;
         L     #S10step;
         T     "Data_to_HNOSS".S10step;
         L     #Sxstep;
         T     "Data_to_HNOSS".SXstep;
END_REGION
END_FUNCTION

FUNCTION "UpdateData2HNOSS" : Void   // FC303, LAD
{ S7_Optimized_Access := 'FALSE' }
AUTHOR : KG
VERSION : 0.1
BEGIN

REGION Network 1: Initial state
